HMI tags "Tank"
   "DB702_Tank_Value.Tank[0].Density" : Int = PLC DB702_Tank_Value.Tank[0].Density AT %DB702.DBW36, 1 s
      on ChangeValue: SetBit("DB702_Tank_Value.Write")
   "DB702_Tank_Value_Tank{0}_Agitator_RunTime" : S5Time = PLC DB702_Tank_Value.Tank[0].Agitator.RunTime AT %DB702.DBW72, 1 s
      on ChangeValue: SetBit("DB702_Tank_Value.Write")
   "DB702_Tank_Value_Tank{0}_Agitator_PauseTime" : S5Time = PLC DB702_Tank_Value.Tank[0].Agitator.PauseTime AT %DB702.DBW74, 1 s
      on ChangeValue: SetBit("DB702_Tank_Value.Write")
   "DB702_Tank_Value_Tank{0}_FillingTimeControl" : S5Time = PLC DB702_Tank_Value.Tank[0].FillingTimeControl AT %DB702.DBW28, 1 s
      on ChangeValue: SetBit("DB702_Tank_Value.Write")
   "Temper_Actual_0" : Int, internal
   "Temper_SetValue_0" : Int AT %DB1.DBW0
   "DB702_Tank_Value.Pt2_Controller[0].Dif_Cooling_ON" : Real = PLC DB702_Tank_Value.Pt2_Controller[0].Dif_Cooling_ON AT %DB702.DBD1072, 1 s
      on ChangeValue: SetBit("DB702_Tank_Value.Write")
   "DB702_Tank_Value.Pt2_Controller[0].Dif_Cooling_OFF" : Real = PLC DB702_Tank_Value.Pt2_Controller[0].Dif_Cooling_OFF AT %DB702.DBD1076, 1 s
      on ChangeValue: SetBit("DB702_Tank_Value.Write")
   "DB702_Tank_Value.Pt2_Controller[0].Dif_Heating_ON" : Real = PLC DB702_Tank_Value.Pt2_Controller[0].Dif_Heating_ON AT %DB702.DBD1080, 1 s
      on ChangeValue: SetBit("DB702_Tank_Value.Write")
   "DB702_Tank_Value.Pt2_Controller[0].Dif_Heating_OFF" : Real = PLC DB702_Tank_Value.Pt2_Controller[0].Dif_Heating_OFF AT %DB702.DBD1084, 1 s
      on ChangeValue: SetBit("DB702_Tank_Value.Write")
   "DB612_Tank_State.Read" : Bool = PLC DB612_Tank_State.Read AT %DB612.DBX6.0, 1 s
   "DB612_Tank_State.Write" : Bool = PLC DB612_Tank_State.Write AT %DB612.DBX6.1, 1 s
   "DB702_Tank_Value.Write" : Bool = PLC DB702_Tank_Value.Write AT %DB702.DBX4.1, 1 s
   "DB612_Tank_State.ActualDeviceNo" : Int = PLC DB612_Tank_State.ActualDeviceNo AT %DB612.DBW2, 1 s
      on ChangeValue: SetBit("DB702_Tank_Value.Write")
   "DB612_Tank_State.ReadDeviceNo" : Int = PLC DB612_Tank_State.ReadDeviceNo AT %DB612.DBW0, 1 s
      on ChangeValue: SetBit("DB702_Tank_Value.Write")
   "DB702_Tank_Value.Tank[0].TankLevel.Max_Level" : Real = PLC DB702_Tank_Value.Tank[0].TankLevel.Max_Level AT %DB702.DBD46, 1 s
      on ChangeValue: SetBit("DB702_Tank_Value.Write")
   "DB702_Tank_Value.Tank[0].TankLevel.Start_Level_Filling" : Real = PLC DB702_Tank_Value.Tank[0].TankLevel.Start_Level_Filling AT %DB702.DBD50, 1 s
      on ChangeValue: SetBit("DB702_Tank_Value.Write")
   "DB702_Tank_Value.Tank[0].TankLevel.Stop_Level_Filling" : Real = PLC DB702_Tank_Value.Tank[0].TankLevel.Stop_Level_Filling AT %DB702.DBD54, 1 s
      on ChangeValue: SetBit("DB702_Tank_Value.Write")
   "DB702_Tank_Value.Tank[0].TankLevel.Stop_Level_Agitator" : Real = PLC DB702_Tank_Value.Tank[0].TankLevel.Stop_Level_Agitator AT %DB702.DBD58, 1 s
      on ChangeValue: SetBit("DB702_Tank_Value.Write")
   "DB702_Tank_Value.Tank[0].TankLevel.Min_Level_Warning" : Real = PLC DB702_Tank_Value.Tank[0].TankLevel.Min_Level_Warning AT %DB702.DBD62, 1 s
      on ChangeValue: SetBit("DB702_Tank_Value.Write")
   "DB702_Tank_Value.Tank[0].TankLevel.Min_Level" : Real = PLC DB702_Tank_Value.Tank[0].TankLevel.Min_Level AT %DB702.DBD66, 1 s
      on ChangeValue: SetBit("DB702_Tank_Value.Write")
   "Open_Tempering_Dialog" : Int, internal
   "Open_Filling_Level_Tank" : Int, internal
   "DB702_Tank_Value_Tank{0}_NoShotFilling" : Int = PLC DB702_Tank_Value.Tank[0].NoShotFilling AT %DB702.DBW30, 1 s
      on ChangeValue: SetBit("DB702_Tank_Value.Write")
   "DB702_Tank_Value_Tank{0}_TimeToStartFilling" : S5Time = PLC DB702_Tank_Value.Tank[0].TimeToStartFilling AT %DB702.DBW32, 1 s
      on ChangeValue: SetBit("DB702_Tank_Value.Write")
   "Tank Load Event" : Int, internal
   "Open_Temperature_Barrel" : Int, internal
   "DB702_Tank_Value_Pt2_ControllerBarell{0}_Dif_Cooling_ON" : Real = PLC DB702_Tank_Value.Pt2_ControllerBarell[0].Dif_Cooling_ON AT %DB702.DBD1384, 1 s
      on ChangeValue: SetBit("DB702_Tank_Value.Write")
   "DB702_Tank_Value_Pt2_ControllerBarell{0}_Dif_Cooling_OFF" : Real = PLC DB702_Tank_Value.Pt2_ControllerBarell[0].Dif_Cooling_OFF AT %DB702.DBD1388, 1 s
      on ChangeValue: SetBit("DB702_Tank_Value.Write")
   "DB702_Tank_Value_Pt2_ControllerBarell{0}_Dif_Heating_ON" : Real = PLC DB702_Tank_Value.Pt2_ControllerBarell[0].Dif_Heating_ON AT %DB702.DBD1392, 1 s
      on ChangeValue: SetBit("DB702_Tank_Value.Write")
   "DB702_Tank_Value_Pt2_ControllerBarell{0}_Dif_Heating_OFF" : Real = PLC DB702_Tank_Value.Pt2_ControllerBarell[0].Dif_Heating_OFF AT %DB702.DBD1396, 1 s
      on ChangeValue: SetBit("DB702_Tank_Value.Write")
   "DB702_Tank_Value_Pt2_ControllerBarell{0}_Max_Temp" : Real = PLC DB702_Tank_Value.Pt2_ControllerBarell[0].Max_Temp AT %DB702.DBD1400, 1 s
      on ChangeValue: SetBit("DB702_Tank_Value.Write")
   "DB702_Tank_Value_Pt2_ControllerBarell{0}_Min_Temp" : Real = PLC DB702_Tank_Value.Pt2_ControllerBarell[0].Min_Temp AT %DB702.DBD1404, 1 s
      on ChangeValue: SetBit("DB702_Tank_Value.Write")
   "DB702_Tank_Value_Tank{0}_With_Vacuum" : Bool = PLC DB702_Tank_Value.Tank[0].With_Vacuum AT %DB702.DBX39.7, 1 s
      on ChangeValue: SetBit("DB702_Tank_Value.Write")
   "DB702_Tank_Value_Tank{0}_With_Nucleation" : Bool = PLC DB702_Tank_Value.Tank[0].With_Nucleation AT %DB702.DBX40.0, 1 s
      on ChangeValue: SetBit("DB702_Tank_Value.Write")
   "DB702_Tank_Value_Tank{0}_Deselected" : Bool = PLC DB702_Tank_Value.Tank[0].Deselected AT %DB702.DBX39.1, 1 s
      on ChangeValue: SetBit("DB702_Tank_Value.Write")
   "DB702_Tank_Value_Tank{0}_With_Filling_Pentane" : Bool = PLC DB702_Tank_Value.Tank[0].With_Filling_Pentane AT %DB702.DBX42.7, 1 s
      on ChangeValue: SetBit("DB702_Tank_Value.Write")
   "DB702_Tank_Value_Tank{0}_Existing" : Bool = PLC DB702_Tank_Value.Tank[0].Existing AT %DB702.DBX39.0, 1 s
      on ChangeValue: SetBit("DB702_Tank_Value.Write")
   "DB702_Tank_Value_Tank{0}_With_Heating" : Bool = PLC DB702_Tank_Value.Tank[0].With_Heating AT %DB702.DBX39.6, 1 s
      on ChangeValue: SetBit("DB702_Tank_Value.Write")
   "DB702_Tank_Value_Tank{0}_With_Filling" : Bool = PLC DB702_Tank_Value.Tank[0].With_Filling AT %DB702.DBX42.0, 1 s
      on ChangeValue: SetBit("DB702_Tank_Value.Write")
   "DB702_Tank_Value_Tank{0}_With_Agitator" : Bool = PLC DB702_Tank_Value.Tank[0].With_Agitator AT %DB702.DBX45.0, 1 s
      on ChangeValue: SetBit("DB702_Tank_Value.Write")
   "DB702_Tank_Value_Tank{0}_With_Agitator_Converter" : Bool = PLC DB702_Tank_Value.Tank[0].With_Agitator_Converter AT %DB702.DBX45.1, 1 s
      on ChangeValue: SetBit("DB702_Tank_Value.Write")
   "DB702_Tank_Value_Tank{0}_With_Agitator_SetValue" : Bool = PLC DB702_Tank_Value.Tank[0].With_Agitator_SetValue AT %DB702.DBX45.2, 1 s
      on ChangeValue: SetBit("DB702_Tank_Value.Write")
   "DB702_Tank_Value_Tank{0}_With_Agitator_6SetValue" : Bool = PLC DB702_Tank_Value.Tank[0].With_Agitator_6SetValue AT %DB702.DBX45.3, 1 s
      on ChangeValue: SetBit("DB702_Tank_Value.Write")
   "DB702_Tank_Value_Tank{0}_With_BarelStation" : Bool = PLC DB702_Tank_Value.Tank[0].With_BarelStation AT %DB702.DBX44.0, 1 s
      on ChangeValue: SetBit("DB702_Tank_Value.Write")
   "DB702_Tank_Value_Tank{0}_With_BarelStation_Zirkulation" : Bool = PLC DB702_Tank_Value.Tank[0].With_BarelStation_Zirkulation AT %DB702.DBX44.1, 1 s
      on ChangeValue: SetBit("DB702_Tank_Value.Write")
   "DB702_Tank_Value_Tank{0}_With_BarelStation_PnPump" : Bool = PLC DB702_Tank_Value.Tank[0].With_BarelStation_PnPump AT %DB702.DBX44.2, 1 s
      on ChangeValue: SetBit("DB702_Tank_Value.Write")
   "DB702_Tank_Value_Tank{0}_With_BarelStation_ElPump" : Bool = PLC DB702_Tank_Value.Tank[0].With_BarelStation_ElPump AT %DB702.DBX44.3, 1 s
      on ChangeValue: SetBit("DB702_Tank_Value.Write")
   "DB702_Tank_Value_Tank{0}_With_BarelStation_PnRW" : Bool = PLC DB702_Tank_Value.Tank[0].With_BarelStation_PnRW AT %DB702.DBX44.4, 1 s
      on ChangeValue: SetBit("DB702_Tank_Value.Write")
   "DB702_Tank_Value_Tank{0}_With_BarelStation_ElRW" : Bool = PLC DB702_Tank_Value.Tank[0].With_BarelStation_ElRW AT %DB702.DBX44.5, 1 s
      on ChangeValue: SetBit("DB702_Tank_Value.Write")
   "DB702_Tank_Value_Tank{0}_With_BarelStation_Heating" : Bool = PLC DB702_Tank_Value.Tank[0].With_BarelStation_Heating AT %DB702.DBX44.6, 1 s
      on ChangeValue: SetBit("DB702_Tank_Value.Write")
   "DB702_Tank_Value_Tank{0}_With_BarelStation_HeatingBottom" : Bool = PLC DB702_Tank_Value.Tank[0].With_BarelStation_HeatingBottom AT %DB702.DBX44.7, 1 s
      on ChangeValue: SetBit("DB702_Tank_Value.Write")
   "DB702_Tank_Value_Tank{0}_With_Tempering" : Bool = PLC DB702_Tank_Value.Tank[0].With_Tempering AT %DB702.DBX43.0, 1 s
      on ChangeValue: SetBit("DB702_Tank_Value.Write")
   "DB702_Tank_Value_Tank{0}_With_Tempering_TempGeraet" : Bool = PLC DB702_Tank_Value.Tank[0].With_Tempering_TempGeraet AT %DB702.DBX43.1, 1 s
      on ChangeValue: SetBit("DB702_Tank_Value.Write")
   "DB702_Tank_Value_Tank{0}_With_Tempering_VKaltwasser" : Bool = PLC DB702_Tank_Value.Tank[0].With_Tempering_VKaltwasser AT %DB702.DBX43.2, 1 s
      on ChangeValue: SetBit("DB702_Tank_Value.Write")
   "DB702_Tank_Value_Tank{0}_With_Tempering_Heizung" : Bool = PLC DB702_Tank_Value.Tank[0].With_Tempering_Heizung AT %DB702.DBX43.3, 1 s
      on ChangeValue: SetBit("DB702_Tank_Value.Write")
   "DB702_Tank_Value_Tank{0}_With_Tempering_WTRL" : Bool = PLC DB702_Tank_Value.Tank[0].With_Tempering_WTRL AT %DB702.DBX43.4, 1 s
      on ChangeValue: SetBit("DB702_Tank_Value.Write")
   "DB702_Tank_Value_Tank{0}_With_Tempering_WTmitFischer" : Bool = PLC DB702_Tank_Value.Tank[0].With_Tempering_WTmitFischer AT %DB702.DBX43.5, 1 s
      on ChangeValue: SetBit("DB702_Tank_Value.Write")
   "DB702_Tank_Value_Tank{0}_With_Tempering_WTBypass" : Bool = PLC DB702_Tank_Value.Tank[0].With_Tempering_WTBypass AT %DB702.DBX43.6, 1 s
      on ChangeValue: SetBit("DB702_Tank_Value.Write")
   "DB702_Tank_Value_Tank{0}_With_Tempering_WTVL" : Bool = PLC DB702_Tank_Value.Tank[0].With_Tempering_WTVL AT %DB702.DBX43.7, 1 s
      on ChangeValue: SetBit("DB702_Tank_Value.Write")
   "DB702_Tank_Value_Tank{0}_With_Filling_Valve" : Bool = PLC DB702_Tank_Value.Tank[0].With_Filling_Valve AT %DB702.DBX42.1, 1 s
      on ChangeValue: SetBit("DB702_Tank_Value.Write")
   "DB702_Tank_Value_Tank{0}_With_Filling_2Valve" : Bool = PLC DB702_Tank_Value.Tank[0].With_Filling_2Valve AT %DB702.DBX42.2, 1 s
      on ChangeValue: SetBit("DB702_Tank_Value.Write")
   "DB702_Tank_Value_Tank{0}_With_Filling_ShutDown" : Bool = PLC DB702_Tank_Value.Tank[0].With_Filling_ShutDown AT %DB702.DBX42.3, 1 s
      on ChangeValue: SetBit("DB702_Tank_Value.Write")
   "DB702_Tank_Value_Tank{0}_With_Filling_Switch" : Bool = PLC DB702_Tank_Value.Tank[0].With_Filling_Switch AT %DB702.DBX42.4, 1 s
      on ChangeValue: SetBit("DB702_Tank_Value.Write")
   "DB702_Tank_Value_Tank{0}_With_Filling_Pump" : Bool = PLC DB702_Tank_Value.Tank[0].With_Filling_Pump AT %DB702.DBX42.5, 1 s
      on ChangeValue: SetBit("DB702_Tank_Value.Write")
   "DB702_Tank_Value_Tank{0}_With_Filling_DryRun" : Bool = PLC DB702_Tank_Value.Tank[0].With_Filling_DryRun AT %DB702.DBX42.6, 1 s
      on ChangeValue: SetBit("DB702_Tank_Value.Write")
   "DB702_Tank_Value_Tank{0}_With_ContainerStation" : Bool = PLC DB702_Tank_Value.Tank[0].With_ContainerStation AT %DB702.DBX40.3, 1 s
      on ChangeValue: SetBit("DB702_Tank_Value.Write")
   "DB702_Tank_Value_Tank{0}_With_Level_3Liq" : Bool = PLC DB702_Tank_Value.Tank[0].With_Level_3Liq AT %DB702.DBX41.0, 1 s
      on ChangeValue: SetBit("DB702_Tank_Value.Write")
   "DB702_Tank_Value_Tank{0}_With_Level_4Liq" : Bool = PLC DB702_Tank_Value.Tank[0].With_Level_4Liq AT %DB702.DBX41.1, 1 s
      on ChangeValue: SetBit("DB702_Tank_Value.Write")
   "DB702_Tank_Value_Tank{0}_With_Level_Probe" : Bool = PLC DB702_Tank_Value.Tank[0].With_Level_Probe AT %DB702.DBX41.2, 1 s
      on ChangeValue: SetBit("DB702_Tank_Value.Write")
   "DB702_Tank_Value_Tank{0}_With_Level_SMin" : Bool = PLC DB702_Tank_Value.Tank[0].With_Level_SMin AT %DB702.DBX41.3, 1 s
      on ChangeValue: SetBit("DB702_Tank_Value.Write")
   "DB702_Tank_Value_Tank{0}_With_Level_SMax" : Bool = PLC DB702_Tank_Value.Tank[0].With_Level_SMax AT %DB702.DBX41.4, 1 s
      on ChangeValue: SetBit("DB702_Tank_Value.Write")
   "DB702_Tank_Value_Tank{0}_With_Triptray" : Bool = PLC DB702_Tank_Value.Tank[0].With_Triptray AT %DB702.DBX41.5, 1 s
      on ChangeValue: SetBit("DB702_Tank_Value.Write")
   "DB702_Tank_Value_Tank{0}_Name" : String[20] = PLC DB702_Tank_Value.Tank[0].Name AT %DB702.DBX6.0, 1 s
      on ChangeValue: SetBit("DB702_Tank_Value.Write")
   "DB702_Tank_Value_Tank{0}_Color" : Byte = PLC DB702_Tank_Value.Tank[0].Color AT %DB702.DBB38, 1 s
      on ChangeValue: SetBit("DB702_Tank_Value.Write")
   "DB702_Tank_Value_Tank{1}_Name" : String[20] = PLC DB702_Tank_Value.Tank[1].Name AT %DB702.DBX82.0, 1 s
      on ChangeValue: SetBit("DB702_Tank_Value.Write")
   "DB702_Tank_Value_Tank{2}_Name" : String[20] = PLC DB702_Tank_Value.Tank[2].Name AT %DB702.DBX158.0, 1 s
      on ChangeValue: SetBit("DB702_Tank_Value.Write")
   "DB702_Tank_Value_Tank{2}_Color" : Byte = PLC DB702_Tank_Value.Tank[2].Color AT %DB702.DBB190, 1 s
      on ChangeValue: SetBit("DB702_Tank_Value.Write")
   "DB702_Tank_Value_Tank{1}_Color" : Byte = PLC DB702_Tank_Value.Tank[1].Color AT %DB702.DBB114, 1 s
      on ChangeValue: SetBit("DB702_Tank_Value.Write")
   "DB702_Tank_Value_Tank{3}_Color" : Byte = PLC DB702_Tank_Value.Tank[3].Color AT %DB702.DBB266, 1 s
      on ChangeValue: SetBit("DB702_Tank_Value.Write")
   "DB702_Tank_Value_Tank{4}_Color" : Byte = PLC DB702_Tank_Value.Tank[4].Color AT %DB702.DBB342, 1 s
      on ChangeValue: SetBit("DB702_Tank_Value.Write")
   "DB702_Tank_Value_Tank{5}_Color" : Byte = PLC DB702_Tank_Value.Tank[5].Color AT %DB702.DBB418, 1 s
      on ChangeValue: SetBit("DB702_Tank_Value.Write")
   "DB702_Tank_Value_Tank{6}_Color" : Byte = PLC DB702_Tank_Value.Tank[6].Color AT %DB702.DBB494, 1 s
      on ChangeValue: SetBit("DB702_Tank_Value.Write")
   "DB702_Tank_Value_CirculationPump{0}_RunTime" : S5Time = PLC DB702_Tank_Value.CirculationPump[0].RunTime AT %DB702.DBW1696, 1 s
   "DB702_Tank_Value_CirculationPump{0}_PauseTime" : S5Time = PLC DB702_Tank_Value.CirculationPump[0].PauseTime AT %DB702.DBW1698, 1 s
   "DB602_PV_Tank_Tank{0}_JacketHeater_PV_ActV_Value" : Real = PLC DB602_PV_Tank.Tank[0].JacketHeater.PV_ActV.Value AT %DB602.DBD218, 1 s
   "DB602_PV_Tank_Tank{0}_JacketHeater_PV_SetV_Value" : Real = PLC DB602_PV_Tank.Tank[0].JacketHeater.PV_SetV.Value AT %DB602.DBD198, 1 s
      on ChangeValue: SetBit("DB702_Tank_Value.Write")
   "DB602_PV_Tank_Tank{0}_Level_PV_SetV_Value" : Real = PLC DB602_PV_Tank.Tank[0].Level.PV_SetV.Value AT %DB602.DBD54, 1 s
      on ChangeValue: SetBit("DB702_Tank_Value.Write")
   "DB602_PV_Tank_Tank{0}_Temp_PV_SetV_Value" : Real = PLC DB602_PV_Tank.Tank[0].Temp.PV_SetV.Value AT %DB602.DBD6, 1 s
      on ChangeValue: SetBit("DB702_Tank_Value.Write")
   "DB602_PV_Tank_Tank{0}_Temp_PV_SetV_WarningLowerLimit" : Real = PLC DB602_PV_Tank.Tank[0].Temp.PV_SetV.WarningLowerLimit AT %DB602.DBD10, 1 s
      on ChangeValue: SetBit("DB702_Tank_Value.Write")
   "DB602_PV_Tank_Tank{0}_Temp_PV_SetV_WarningUpperLimit" : Real = PLC DB602_PV_Tank.Tank[0].Temp.PV_SetV.WarningUpperLimit AT %DB602.DBD14, 1 s
      on ChangeValue: SetBit("DB702_Tank_Value.Write")
   "DB602_PV_Tank_Tank{0}_Temp_PV_SetV_AlarmLowerLimit" : Real = PLC DB602_PV_Tank.Tank[0].Temp.PV_SetV.AlarmLowerLimit AT %DB602.DBD18, 1 s
      on ChangeValue: SetBit("DB702_Tank_Value.Write")
   "DB602_PV_Tank_Tank{0}_Temp_PV_SetV_AlarmUpperLimit" : Real = PLC DB602_PV_Tank.Tank[0].Temp.PV_SetV.AlarmUpperLimit AT %DB602.DBD22, 1 s
      on ChangeValue: SetBit("DB702_Tank_Value.Write")
   "DB602_PV_Tank_Tank{0}_Nucleation_PV_SetV_Value" : Real = PLC DB602_PV_Tank.Tank[0].Nucleation.PV_SetV.Value AT %DB602.DBD150, 1 s
      on ChangeValue: SetBit("DB702_Tank_Value.Write")
   "DB602_PV_Tank_Tank{0}_Nucleation_PV_SetV_WarningLowerLimit" : Real = PLC DB602_PV_Tank.Tank[0].Nucleation.PV_SetV.WarningLowerLimit AT %DB602.DBD154, 1 s
      on ChangeValue: SetBit("DB702_Tank_Value.Write")
   "DB602_PV_Tank_Tank{0}_Nucleation_PV_SetV_WarningUpperLimit" : Real = PLC DB602_PV_Tank.Tank[0].Nucleation.PV_SetV.WarningUpperLimit AT %DB602.DBD158, 1 s
      on ChangeValue: SetBit("DB702_Tank_Value.Write")
   "DB602_PV_Tank_Tank{0}_Nucleation_PV_SetV_AlarmLowerLimit" : Real = PLC DB602_PV_Tank.Tank[0].Nucleation.PV_SetV.AlarmLowerLimit AT %DB602.DBD162, 1 s
      on ChangeValue: SetBit("DB702_Tank_Value.Write")
   "DB602_PV_Tank_Tank{0}_Nucleation_PV_SetV_AlarmUpperLimit" : Real = PLC DB602_PV_Tank.Tank[0].Nucleation.PV_SetV.AlarmUpperLimit AT %DB602.DBD166, 1 s
      on ChangeValue: SetBit("DB702_Tank_Value.Write")
   "DB612_Tank_State_Tank{0}_Switch_Refilling_from_Barrel_ON_OFF" : Bool = PLC DB612_Tank_State.Tank[0].Switch_Refilling_from_Barrel_ON_OFF AT %DB612.DBX15.3, 1 s
      on ChangeValue: SetBit("DB612_Tank_State.Write")
   "DB612_Tank_State_ControllerTankTemp{0}_Switch_Temp_ON_OFF" : Bool = PLC DB612_Tank_State.ControllerTankTemp[0].Switch_Temp_ON_OFF AT %DB612.DBX375.7, 1 s
      on ChangeValue: SetBit("DB612_Tank_State.Write")
   "DB612_Tank_State_Tank{0}_Switch_Refilling_ON_OFF" : Bool = PLC DB612_Tank_State.Tank[0].Switch_Refilling_ON_OFF AT %DB612.DBX14.6, 1 s
      on ChangeValue: SetBit("DB612_Tank_State.Write")
   "DB612_Tank_State_ControllerBarellTemp{0}_Switch_Temp_ON_OFF" : Bool = PLC DB612_Tank_State.ControllerBarellTemp[0].Switch_Temp_ON_OFF AT %DB612.DBX583.7, 1 s
      on ChangeValue: SetBit("DB612_Tank_State.Write")
   "DB612_Tank_State_Vacuum{0}_Switch_Vacuum_ON_OFF" : Bool = PLC DB612_Tank_State.Vacuum[0].Switch_Vacuum_ON_OFF AT %DB612.DBX218.2, 1 s
      on ChangeValue: SetBit("DB612_Tank_State.Write")
   "DB612_Tank_State_CirculationPump{0}_Switch_Drive_ON_OFF" : Bool = PLC DB612_Tank_State.CirculationPump[0].Switch_Drive_ON_OFF AT %DB612.DBX271.7, 1 s
      on ChangeValue: SetBit("DB612_Tank_State.Write")
   "DB612_Tank_State_Tank{0}_Switch_DrainTank_ON_OFF" : Bool = PLC DB612_Tank_State.Tank[0].Switch_DrainTank_ON_OFF AT %DB612.DBX15.1, 1 s
      on ChangeValue: SetBit("DB612_Tank_State.Write")
   "DB612_Tank_State_Agitator{0}_Switch_Drive_ON_OFF" : Bool = PLC DB612_Tank_State.Agitator[0].Switch_Drive_ON_OFF AT %DB612.DBX115.6, 1 s
      on ChangeValue: SetBit("DB612_Tank_State.Write")
   "DB612_Tank_State_FaultExists{1}" : Bool = PLC DB612_Tank_State.FaultExists[1] AT %DB612.DBX8.1, 1 s
   "DB612_Tank_State_FaultExists{2}" : Bool = PLC DB612_Tank_State.FaultExists[2] AT %DB612.DBX8.2, 1 s
   "DB612_Tank_State_Tank{0}_State_Refilling" : Int = PLC DB612_Tank_State.Tank[0].State_Refilling AT %DB612.DBW16, 1 s
   "DB702_Tank_Value_Tank{0}_With_Drain" : Bool = PLC DB702_Tank_Value.Tank[0].With_Drain AT %DB702.DBX40.2, 1 s
      on ChangeValue: SetBit("DB702_Tank_Value.Write")
   "DB702_Tank_Value_Tank{0}_Agitator_Config_bit_Heating_ON" : Bool = PLC DB702_Tank_Value.Tank[0].Agitator.Config_bit_Heating_ON AT %DB702.DBX70.2, 1 s
      on ChangeValue: SetBit("DB702_Tank_Value.Write")
   "DB702_Tank_Value_Tank{0}_Agitator_Config_bit_Cooling_ON" : Bool = PLC DB702_Tank_Value.Tank[0].Agitator.Config_bit_Cooling_ON AT %DB702.DBX70.4, 1 s
      on ChangeValue: SetBit("DB702_Tank_Value.Write")
   "DB702_Tank_Value_Tank{0}_Agitator_Config_bit_Filling_ON" : Bool = PLC DB702_Tank_Value.Tank[0].Agitator.Config_bit_Filling_ON AT %DB702.DBX70.6, 1 s
      on ChangeValue: SetBit("DB702_Tank_Value.Write")
   "DB702_Tank_Value_Tank{0}_Agitator_config_bit_Heating_Int" : Bool = PLC DB702_Tank_Value.Tank[0].Agitator.config_bit_Heating_Int AT %DB702.DBX70.3, 1 s
      on ChangeValue: SetBit("DB702_Tank_Value.Write")
   "DB702_Tank_Value_Tank{0}_Agitator_Config_bit_Cooling_Int" : Bool = PLC DB702_Tank_Value.Tank[0].Agitator.Config_bit_Cooling_Int AT %DB702.DBX70.5, 1 s
      on ChangeValue: SetBit("DB702_Tank_Value.Write")
   "DB702_Tank_Value_Tank{0}_Agitator_Config_bit_Filling_Int" : Bool = PLC DB702_Tank_Value.Tank[0].Agitator.Config_bit_Filling_Int AT %DB702.DBX70.7, 1 s
      on ChangeValue: SetBit("DB702_Tank_Value.Write")
   "DB702_Tank_Value_Tank{0}_Agitator_Config_bit_Charging_ON" : Bool = PLC DB702_Tank_Value.Tank[0].Agitator.Config_bit_Charging_ON AT %DB702.DBX71.0, 1 s
      on ChangeValue: SetBit("DB702_Tank_Value.Write")
   "DB702_Tank_Value_Tank{0}_Agitator_Config_bit_Charging_Int" : Bool = PLC DB702_Tank_Value.Tank[0].Agitator.Config_bit_Charging_Int AT %DB702.DBX71.1, 1 s
      on ChangeValue: SetBit("DB702_Tank_Value.Write")
   "DB702_Tank_Value_Tank{0}_Agitator_Config_bit_Converter" : Bool = PLC DB702_Tank_Value.Tank[0].Agitator.Config_bit_Converter AT %DB702.DBX70.0, 1 s
      on ChangeValue: SetBit("DB702_Tank_Value.Write")
   "DB702_Tank_Value_Tank{0}_With_Level" : Bool = PLC DB702_Tank_Value.Tank[0].With_Level AT %DB702.DBX39.3, 1 s
      on ChangeValue: SetBit("DB702_Tank_Value.Write")
   "DB702_Tank_Value_Tank{0}_PreAgitatingTime" : S5Time = PLC DB702_Tank_Value.Tank[0].PreAgitatingTime AT %DB702.DBW34, 1 s
      on ChangeValue: SetBit("DB702_Tank_Value.Write")
   "DB612_Tank_State_Agitator{0}_State_Drive" : Int = PLC DB612_Tank_State.Agitator[0].State_Drive AT %DB612.DBW116, 1 s
   "DB612_Tank_State_ControllerTankTemp{0}_State_Temp" : Int = PLC DB612_Tank_State.ControllerTankTemp[0].State_Temp AT %DB612.DBW380, 1 s
   "DB612_Tank_State_ControllerBarellTemp{0}_State_Temp" : Int = PLC DB612_Tank_State.ControllerBarellTemp[0].State_Temp AT %DB612.DBW588, 1 s
   "DB612_Tank_State_CirculationPump{0}_State_Drive" : Int = PLC DB612_Tank_State.CirculationPump[0].State_Drive AT %DB612.DBW272, 1 s
   "DB612_Tank_State_Vacuum{0}_Status_Vacuum" : Int = PLC DB612_Tank_State.Vacuum[0].Status_Vacuum AT %DB612.DBW220, 1 s
   "DB702_Tank_Value_Tank{1}_With_Agitator" : Bool = PLC DB702_Tank_Value.Tank[1].With_Agitator AT %DB702.DBX121.0, 1 s
   "DB702_Tank_Value_Tank{2}_With_Agitator" : Bool = PLC DB702_Tank_Value.Tank[2].With_Agitator AT %DB702.DBX197.0, 1 s
   "DB612_Tank_State_Tank{0}_Fault_Exist" : Bool = PLC DB612_Tank_State.Tank[0].Fault_Exist AT %DB612.DBX12.0, 1 s
   "DB612_Tank_State_FaulExist" : Bool = PLC DB612_Tank_State.FaulExist AT %DB612.DBX6.3, 1 s
   "DB612_Tank_State_Agitator{0}_FLT_Exist" : Bool = PLC DB612_Tank_State.Agitator[0].FLT_Exist AT %DB612.DBX114.0, 1 s
   "DB612_Tank_State_AgitatorBarell{0}_FLT_Exist" : Bool = PLC DB612_Tank_State.AgitatorBarell[0].FLT_Exist AT %DB612.DBX166.0, 1 s
   "DB612_Tank_State_Vacuum{0}_FLT_PVacuum" : Bool = PLC DB612_Tank_State.Vacuum[0].FLT_PVacuum AT %DB612.DBX219.0, 1 s
   "DB612_Tank_State_CirculationPump{0}_FaultExist" : Bool = PLC DB612_Tank_State.CirculationPump[0].FaultExist AT %DB612.DBX270.7, 1 s
   "DB612_Tank_State_Pentan{0}_Fault_Exist" : Bool = PLC DB612_Tank_State.Pentan[0].Fault_Exist AT %DB612.DBX348.0, 1 s
   "DB612_Tank_State_ControllerTankTemp{0}_Fault_Exist" : Bool = PLC DB612_Tank_State.ControllerTankTemp[0].Fault_Exist AT %DB612.DBX375.2, 1 s
   "DB612_Tank_State_ControllerTankJacketHeater{0}_Fault_Exist" : Bool = PLC DB612_Tank_State.ControllerTankJacketHeater[0].Fault_Exist AT %DB612.DBX479.2, 1 s
   "DB612_Tank_State_ControllerBarellTemp{0}_Fault_Exist" : Bool = PLC DB612_Tank_State.ControllerBarellTemp[0].Fault_Exist AT %DB612.DBX583.2, 1 s
   "DB612_Tank_State_Tank{0}_Max_Level" : Bool = PLC DB612_Tank_State.Tank[0].Max_Level AT %DB612.DBX14.1, 1 s
   "DB612_Tank_State_Tank{0}_Min_Level" : Bool = PLC DB612_Tank_State.Tank[0].Min_Level AT %DB612.DBX14.4, 1 s
   "DB612_Tank_State_Tank{0}_Filling_Start" : Bool = PLC DB612_Tank_State.Tank[0].Filling_Start AT %DB612.DBX13.5, 1 s
   "DB612_Tank_State_Tank{0}_Stop_Level_Filling" : Bool = PLC DB612_Tank_State.Tank[0].Stop_Level_Filling AT %DB612.DBX14.2, 1 s
   "DB612_Tank_State_Tank{0}_Start_Level_Filling" : Bool = PLC DB612_Tank_State.Tank[0].Start_Level_Filling AT %DB612.DBX14.3, 1 s
   "DB702_Tank_Value_Tank{2}_With_Filling" : Bool = PLC DB702_Tank_Value.Tank[2].With_Filling AT %DB702.DBX194.0, 1 s
   "DB702_Tank_Value_Tank{1}_With_Filling" : Bool = PLC DB702_Tank_Value.Tank[1].With_Filling AT %DB702.DBX118.0, 1 s
   "DB702_Tank_Value_Tank{1}_With_Tempering_Heizung" : Bool = PLC DB702_Tank_Value.Tank[1].With_Tempering_Heizung AT %DB702.DBX119.3, 1 s
   "DB702_Tank_Value_Tank{2}_With_Tempering_Heizung" : Bool = PLC DB702_Tank_Value.Tank[2].With_Tempering_Heizung AT %DB702.DBX195.3, 1 s
   "DB702_Tank_Value_Tank{3}_Name" : String[20] = PLC DB702_Tank_Value.Tank[3].Name AT %DB702.DBX234.0, 1 s
   "DB702_Tank_Value_Tank{4}_Name" : String[20] = PLC DB702_Tank_Value.Tank[4].Name AT %DB702.DBX310.0, 1 s
   "DB702_Tank_Value_Tank{5}_Name" : String[20] = PLC DB702_Tank_Value.Tank[5].Name AT %DB702.DBX386.0, 1 s
   "DB702_Tank_Value_Tank{6}_Name" : String[20] = PLC DB702_Tank_Value.Tank[6].Name AT %DB702.DBX462.0, 1 s
   "DB702_Tank_Value_Tank{7}_Name" : String[20] = PLC DB702_Tank_Value.Tank[7].Name AT %DB702.DBX538.0, 1 s
   "DB702_Tank_Value_Tank{8}_Name" : String[20] = PLC DB702_Tank_Value.Tank[8].Name AT %DB702.DBX614.0, 1 s
   "DB702_Tank_Value_Tank{9}_Name" : String[20] = PLC DB702_Tank_Value.Tank[9].Name AT %DB702.DBX690.0, 1 s
   "DB702_Tank_Value_Tank{10}_Name" : String[20] = PLC DB702_Tank_Value.Tank[10].Name AT %DB702.DBX766.0, 1 s
   "DB702_Tank_Value_Tank{11}_Name" : String[20] = PLC DB702_Tank_Value.Tank[11].Name AT %DB702.DBX842.0, 1 s
   "DB702_Tank_Value_Tank{12}_Name" : String[20] = PLC DB702_Tank_Value.Tank[12].Name AT %DB702.DBX918.0, 1 s
   "DB702_Tank_Value_Tank{1}_With_Level_Probe" : Bool = PLC DB702_Tank_Value.Tank[1].With_Level_Probe AT %DB702.DBX117.2, 1 s
   "DB702_Tank_Value_Tank{2}_With_Level_Probe" : Bool = PLC DB702_Tank_Value.Tank[2].With_Level_Probe AT %DB702.DBX193.2, 1 s
   "DB612_Tank_State_Agitator{0}_Run" : Bool = PLC DB612_Tank_State.Agitator[0].Run AT %DB612.DBX115.0, 1 s
   "DB612_Tank_State_Tank{1}_Start_Level_Filling" : Bool = PLC DB612_Tank_State.Tank[1].Start_Level_Filling AT %DB612.DBX22.3, 1 s
   "DB612_Tank_State_Tank{2}_Start_Level_Filling" : Bool = PLC DB612_Tank_State.Tank[2].Start_Level_Filling AT %DB612.DBX30.3, 1 s
   "DB612_Tank_State_Tank{1}_Stop_Level_Filling" : Bool = PLC DB612_Tank_State.Tank[1].Stop_Level_Filling AT %DB612.DBX22.2, 1 s
   "DB612_Tank_State_Tank{2}_Stop_Level_Filling" : Bool = PLC DB612_Tank_State.Tank[2].Stop_Level_Filling AT %DB612.DBX30.2, 1 s
   "DB612_Tank_State_Tank{2}_Max_Level" : Bool = PLC DB612_Tank_State.Tank[2].Max_Level AT %DB612.DBX30.1, 1 s
   "DB612_Tank_State_Tank{1}_Max_Level" : Bool = PLC DB612_Tank_State.Tank[1].Max_Level AT %DB612.DBX22.1, 1 s
   "DB612_Tank_State_Tank{1}_Min_Level" : Bool = PLC DB612_Tank_State.Tank[1].Min_Level AT %DB612.DBX22.4, 1 s
   "DB612_Tank_State_Tank{2}_Min_Level" : Bool = PLC DB612_Tank_State.Tank[2].Min_Level AT %DB612.DBX30.4, 1 s

HMI tags "Selector"
   "Switch1" : Int, internal
   "DB611_Hydraulic_State_MH_Hydraulic{0}_Switch_Hydraulic_ON_OFF" : Bool = PLC DB611_Hydraulic_State.MH_Hydraulic[0].Switch_Hydraulic_ON_OFF AT %DB611.DBX10.3, 1 s
   "DB619_State_MPart_Recirculation{0}_Intervall" : Bool = PLC DB619_State_MPart.Recirculation[0].Intervall AT %DB619.DBX14.0, 1 s
   "DB619_State_MPart_Recirculation{0}_Lowpressure" : Bool = PLC DB619_State_MPart.Recirculation[0].Lowpressure AT %DB619.DBX14.2, 1 s
   "DB619_State_MPart_Recirculation{0}_Reduced" : Bool = PLC DB619_State_MPart.Recirculation[0].Reduced AT %DB619.DBX14.3, 1 s
   "DB612_Tank_State_ControllerTankTemp{1}_Switch_Temp_ON_OFF" : Bool = PLC DB612_Tank_State.ControllerTankTemp[1].Switch_Temp_ON_OFF AT %DB612.DBX383.7, 1 s
   "DB612_Tank_State_Tank{1}_Switch_Refilling_ON_OFF" : Bool = PLC DB612_Tank_State.Tank[1].Switch_Refilling_ON_OFF AT %DB612.DBX22.6, 1 s
   "DB612_Tank_State_Agitator{1}_Switch_Drive_ON_OFF" : Bool = PLC DB612_Tank_State.Agitator[1].Switch_Drive_ON_OFF AT %DB612.DBX119.6, 1 s
   "DB612_Tank_State_Agitator{2}_Switch_Drive_ON_OFF" : Bool = PLC DB612_Tank_State.Agitator[2].Switch_Drive_ON_OFF AT %DB612.DBX123.6, 1 s
   "DB612_Tank_State_ControllerTankTemp{2}_Switch_Temp_ON_OFF" : Bool = PLC DB612_Tank_State.ControllerTankTemp[2].Switch_Temp_ON_OFF AT %DB612.DBX391.7, 1 s
   "DB612_Tank_State_Tank{2}_Switch_Refilling_ON_OFF" : Bool = PLC DB612_Tank_State.Tank[2].Switch_Refilling_ON_OFF AT %DB612.DBX30.6, 1 s
   "DB613_Komponent_State_EdgeFilter{1}_Switch_Drive_ON_OFF" : Bool = PLC DB613_Komponent_State.EdgeFilter[1].Switch_Drive_ON_OFF AT %DB613.DBX13.7, 1 s
   "DB613_Komponent_State_HeatexchangerLP{1}_Switch_Temp_ON_OFF" : Bool = PLC DB613_Komponent_State.HeatexchangerLP[1].Switch_Temp_ON_OFF AT %DB613.DBX875.7, 1 s
   "DB613_Komponent_State_EdgeFilter{2}_Switch_Drive_ON_OFF" : Bool = PLC DB613_Komponent_State.EdgeFilter[2].Switch_Drive_ON_OFF AT %DB613.DBX17.7, 1 s
   "DB14_TP_Shortcuts_TP_Shortcuts_ButtonNo_4" : Bool = PLC DB14_TP_Shortcuts.TP_Shortcuts.ButtonNo.4, 1 s
   "DB611_Hydraulic_State_MH_Hydraulic{0}_State_Hydraulic" : Int = PLC DB611_Hydraulic_State.MH_Hydraulic[0].State_Hydraulic AT %DB611.DBW12, 1 s
   "DB611_Hydraulic_State_MH_Hydraulic{1}_State_Hydraulic" : Int = PLC DB611_Hydraulic_State.MH_Hydraulic[1].State_Hydraulic AT %DB611.DBW20, 1 s
   "DB611_Hydraulic_State_MH_Hydraulic{1}_Switch_Hydraulic_ON_OFF" : Bool = PLC DB611_Hydraulic_State.MH_Hydraulic[1].Switch_Hydraulic_ON_OFF AT %DB611.DBX18.3, 1 s
   "DB619_State_MPart_Recirculation{0}_State_Intervall" : Int = PLC DB619_State_MPart.Recirculation[0].State_Intervall AT %DB619.DBW18, 1 s
   "DB619_State_MPart_Recirculation{0}_State_Lowpressure" : Int = PLC DB619_State_MPart.Recirculation[0].State_Lowpressure AT %DB619.DBW20, 1 s
   "DB619_State_MPart_Recirculation{0}_State_Reduced" : Int = PLC DB619_State_MPart.Recirculation[0].State_Reduced AT %DB619.DBW22, 1 s
   "DB612_Tank_State_Tank{1}_State_Refilling" : Int = PLC DB612_Tank_State.Tank[1].State_Refilling AT %DB612.DBW24, 1 s
   "DB612_Tank_State_ControllerTankTemp{1}_State_Temp" : Int = PLC DB612_Tank_State.ControllerTankTemp[1].State_Temp AT %DB612.DBW388, 1 s
   "DB612_Tank_State_ControllerTankTemp{2}_State_Temp" : Int = PLC DB612_Tank_State.ControllerTankTemp[2].State_Temp AT %DB612.DBW396, 1 s
   "DB612_Tank_State_Tank{2}_State_Refilling" : Int = PLC DB612_Tank_State.Tank[2].State_Refilling AT %DB612.DBW32, 1 s
   "DB612_Tank_State_Agitator{1}_State_Drive" : Int = PLC DB612_Tank_State.Agitator[1].State_Drive AT %DB612.DBW120, 1 s
   "DB612_Tank_State_Agitator{2}_State_Drive" : Int = PLC DB612_Tank_State.Agitator[2].State_Drive AT %DB612.DBW124, 1 s
   "DB613_Komponent_State_EdgeFilter{1}_State_Drive" : Int = PLC DB613_Komponent_State.EdgeFilter[1].State_Drive AT %DB613.DBW14, 1 s
   "DB613_Komponent_State_EdgeFilter{2}_State_Drive" : Int = PLC DB613_Komponent_State.EdgeFilter[2].State_Drive AT %DB613.DBW18, 1 s
   "DB613_Komponent_State_HeatexchangerLP{2}_Switch_Temp_ON_OFF" : Bool = PLC DB613_Komponent_State.HeatexchangerLP[2].Switch_Temp_ON_OFF AT %DB613.DBX883.7, 1 s
   "DB613_Komponent_State_HeatexchangerLP{2}_State_Temp" : Int = PLC DB613_Komponent_State.HeatexchangerLP[2].State_Temp AT %DB613.DBW888, 1 s
   "DB613_Komponent_State_HeatexchangerLP{1}_State_Temp" : Int = PLC DB613_Komponent_State.HeatexchangerLP[1].State_Temp AT %DB613.DBW880, 1 s
   "DB613_Komponent_State_HeatexchangerHP{1}_Switch_Temp_ON_OFF" : Bool = PLC DB613_Komponent_State.HeatexchangerHP[1].Switch_Temp_ON_OFF AT %DB613.DBX771.7, 1 s
   "DB613_Komponent_State_HeatexchangerHP{1}_State_Temp" : Int = PLC DB613_Komponent_State.HeatexchangerHP[1].State_Temp AT %DB613.DBW776, 1 s
   "DB613_Komponent_State_HeatexchangerHP{2}_Switch_Temp_ON_OFF" : Bool = PLC DB613_Komponent_State.HeatexchangerHP[2].Switch_Temp_ON_OFF AT %DB613.DBX779.7, 1 s
   "DB613_Komponent_State_HeatexchangerHP{2}_State_Temp" : Int = PLC DB613_Komponent_State.HeatexchangerHP[2].State_Temp AT %DB613.DBW784, 1 s
   "DB619_State_MPart_Recirculation{1}_State_Reduced" : Int = PLC DB619_State_MPart.Recirculation[1].State_Reduced AT %DB619.DBW50, 1 s
   "DB619_State_MPart_Recirculation{1}_State_Lowpressure" : Int = PLC DB619_State_MPart.Recirculation[1].State_Lowpressure AT %DB619.DBW48, 1 s
   "DB619_State_MPart_Recirculation{1}_State_Intervall" : Int = PLC DB619_State_MPart.Recirculation[1].State_Intervall AT %DB619.DBW46, 1 s
   "DB611_Hydraulic_State_MH_Hydraulic{2}_State_Hydraulic" : Int = PLC DB611_Hydraulic_State.MH_Hydraulic[2].State_Hydraulic AT %DB611.DBW28, 1 s